REGION Network 8: End Switch
   #tmON_WaitReopenConn(IN := #tPhases.xReopenConnection, PT := T#1s);   // TON
   #tPhases.xEndSwitch := #tmON_WaitReopenConn.Q;
   IF #tmON_WaitReopenConn.Q THEN #tPhases.xReopenConnection := FALSE; END_IF;
END_REGION

REGION Network 9: - - - - - - - - Send - - - - - - - - -
END_REGION

REGION Network 10: Send Data Time Out
   #tmON_TimeoutSendData(IN := #tPhases.xRequestSend, PT := #CONST_DTIMEOUTSENDDATA_MS);   // TON
END_REGION

REGION Network 11: Request Send
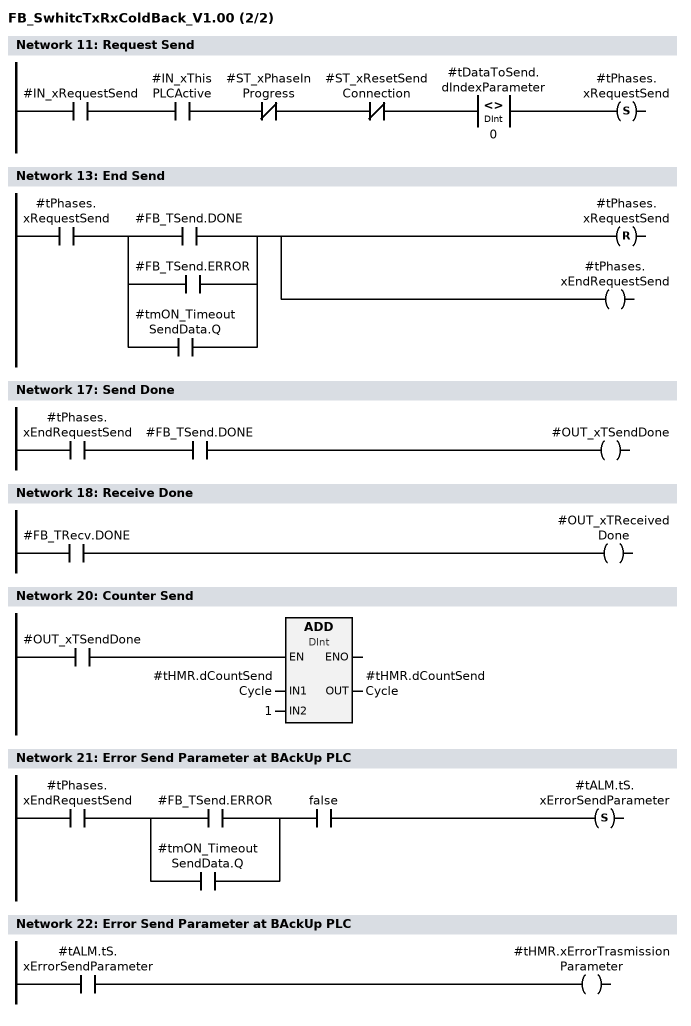
   RUNG wire#powerrail
      Contact( #IN_xRequestSend )
      Contact( #IN_xThisPLCActive )
      I_Contact( #ST_xPhaseInProgress )
      I_Contact( #ST_xResetSendConnection )
      { S7_Templates := "SrcType := DInt" } NE_Contact(in1 := #tDataToSend.dIndexParameter, in2 := 0)
      S_Coil( #tPhases.xRequestSend )
   END_RUNG
   // the same network as SCL:
   IF #IN_xRequestSend AND #IN_xThisPLCActive AND NOT #ST_xPhaseInProgress AND NOT #ST_xResetSendConnection AND (#tDataToSend.dIndexParameter <> 0) THEN
       #tPhases.xRequestSend := TRUE;
   END_IF;
END_REGION

REGION Network 12 (SCL): Send Function
       #AUX_dNumByteToSend := #tDataToSend.dByteToSend+8;//(byte for the index to send and the byte so send
   IF #tPhases.xCloseExistinConnection OR NOT #ST_xPLCActive THEN
       #FB_TSend(REQ :=FALSE,
                 CONT := FALSE,
                 LEN := #AUX_dNumByteToSend,
                 CONNECT := #AUX_tConnDataTSend,
                 DATA := #tDataToSend,
                 COM_RST := #ST_xResetSendConnection);

   ELSE
       #FB_TSend(REQ := #tPhases.xRequestSend,
                 CONT := true,
                 LEN := #AUX_dNumByteToSend,
                 CONNECT := #AUX_tConnDataTSend,
                 DATA := #tDataToSend,
                 COM_RST := #ST_xResetSendConnection);
   END_IF;
END_REGION

REGION Network 13: End Send
   RUNG wire#powerrail
      Contact( #tPhases.xRequestSend )
      wire#w1
      Contact( #FB_TSend.DONE )
      wire#w2
      R_Coil( #tPhases.xRequestSend )
   END_RUNG
   RUNG wire#w1
      Contact( #FB_TSend.ERROR )
   END_RUNG wire#w2
   RUNG wire#w1
      Contact( #tmON_TimeoutSendData.Q )
   END_RUNG wire#w2
   RUNG wire#w2
      Coil( #tPhases.xEndRequestSend )
   END_RUNG
   // the same network as SCL:
   #_w1 := #tPhases.xRequestSend AND (#FB_TSend.DONE OR #FB_TSend.ERROR OR #tmON_TimeoutSendData.Q);
   IF #_w1 THEN #tPhases.xRequestSend := FALSE; END_IF;
   #tPhases.xEndRequestSend := #_w1;
END_REGION

REGION Network 14: - - - - - - - - Recive - - - - - - - - -
END_REGION

REGION Network 15 (SCL): Recived Connection
   IF #tPhases.xCloseExistinConnection OR  #ST_xPLCActive THEN
       #FB_TRecv(EN_R := FALSE,
                 CONT := FALSE,
                 LEN := 0,
                 ADHOC:=TRUE,
                 CONNECT := #AUX_tConnDataTRecive,
                 DATA := #tDataRecived,
                 COM_RST := #ST_xResetRecvConnection);
   ELSE
       //Clean DB data recive
       FILL_BLK(IN := 0,
                COUNT := 501,
                OUT => #tDataRecived.rgbSendBuffer[0]);

       #FB_TRecv(EN_R := True,
                  CONT := True,
                  LEN := 0,
                  ADHOC:=TRUE,
                  CONNECT := #AUX_tConnDataTRecive,
                  DATA := #tDataRecived,
                  COM_RST := #ST_xResetRecvConnection);
   END_IF;
END_REGION

REGION Network 16 (SCL): Phase in progress
   GATHER(IN:=#tPhases,
          OUT=>#TMP_dwValue);

   IF #TMP_dwValue <> 0 THEN
       #ST_xPhaseInProgress := TRUE;
   ELSE
       #ST_xPhaseInProgress := FALSE;
   END_IF;
END_REGION

REGION Network 17: Send Done
   RUNG wire#powerrail
      Contact( #tPhases.xEndRequestSend )
      Contact( #FB_TSend.DONE )
      Coil( #OUT_xTSendDone )
   END_RUNG
   // the same network as SCL:
   #OUT_xTSendDone := #tPhases.xEndRequestSend AND #FB_TSend.DONE;
END_REGION

REGION Network 18: Receive Done
   RUNG wire#powerrail
      Contact( #FB_TRecv.DONE )
      Coil( #OUT_xTReceivedDone )
   END_RUNG
   // the same network as SCL:
   #OUT_xTReceivedDone := #FB_TRecv.DONE;
END_REGION

REGION Network 19: - - - - - - - -- - - HMI - - - - - - -
END_REGION

REGION Network 20: Counter Send
   RUNG wire#powerrail
      Contact( #OUT_xTSendDone )
      { S7_Templates := "SrcType := DInt" } Add(in1 := #tHMR.dCountSendCycle, in2 := 1, out => #tHMR.dCountSendCycle)
   END_RUNG
   // the same network as SCL:
   IF #OUT_xTSendDone THEN #tHMR.dCountSendCycle := #tHMR.dCountSendCycle + 1; END_IF;
END_REGION

REGION Network 21: Error Send Parameter at BAckUp PLC
   RUNG wire#powerrail
      Contact( #tPhases.xEndRequestSend )
      wire#w1
      Contact( #FB_TSend.ERROR )
      wire#w2
      Contact( false )
      S_Coil( #tALM.tS.xErrorSendParameter )
   END_RUNG
   RUNG wire#w1
      Contact( #tmON_TimeoutSendData.Q )
   END_RUNG wire#w2
   // the same network as SCL:
   IF #tPhases.xEndRequestSend AND (#FB_TSend.ERROR OR #tmON_TimeoutSendData.Q) AND false THEN
       #tALM.tS.xErrorSendParameter := TRUE;
   END_IF;
END_REGION

REGION Network 22: Error Send Parameter at BAckUp PLC
   RUNG wire#powerrail
      Contact( #tALM.tS.xErrorSendParameter )
      Coil( #tHMR.xErrorTrasmissionParameter )
   END_RUNG
   // the same network as SCL:
   #tHMR.xErrorTrasmissionParameter := #tALM.tS.xErrorSendParameter;
END_REGION
END_FUNCTION_BLOCK

FUNCTION "ExChangeParTxRx_Logic" : Void   // FC340, LAD
{ S7_Optimized_Access := 'TRUE' }
VERSION : 0.1
   VAR_INPUT
      IN_tConfDataMaster : Struct   // Configuration data master CPU
         Header : IF_CONF_Header;
         IPData : IF_CONF_v4;
         NoS : IF_CONF_NOS;
         NTP : IF_CONF_NTP;
         IP_V6 : IF_CONF_v6;
         MAC : IF_CONF_MAC;
         DNS : IF_CONF_DNS;
      END_STRUCT;
      IN_tConfDataBackup : Struct   // Configuration data backup CPU
         Header : IF_CONF_Header;
         IPData : IF_CONF_v4;
         NoS : IF_CONF_NOS;
         NTP : IF_CONF_NTP;
         IP_V6 : IF_CONF_v6;
         MAC : IF_CONF_MAC;
         DNS : IF_CONF_DNS;
      END_STRUCT;
   END_VAR
   VAR_TEMP
      TMP_x : Bool;
      TMP_dBufferPos : DInt;
      TMP_xRetValue : Int;
      IpAddress : IP_V4;
   END_VAR
BEGIN

REGION Network 1 (SCL): IP Secondary CPU
   #IpAddress.ADDR[1] := 192;
   #IpAddress.ADDR[2] := 168;
   #IpAddress.ADDR[3] := 130;
   #IpAddress.ADDR[4] := 8;
END_REGION

REGION Network 2: Call Function Swtich Send/Recive
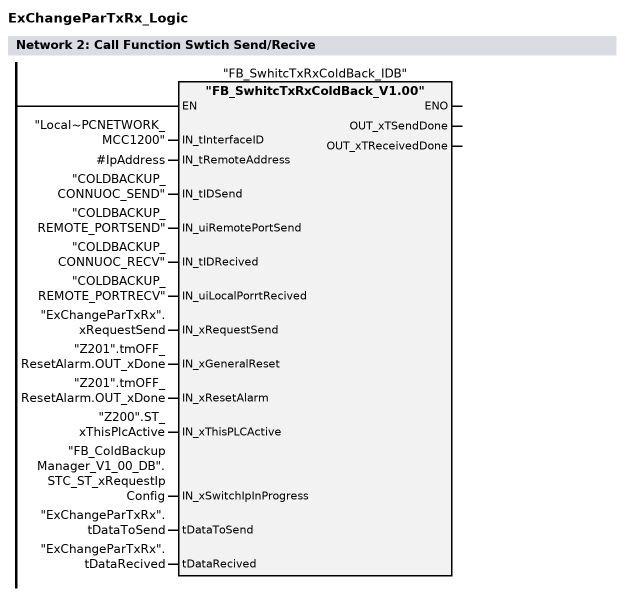
   RUNG wire#powerrail
      "FB_SwhitcTxRxColdBack_IDB"(IN_tInterfaceID := "Local~PCNETWORK_MCC1200", IN_tRemoteAddress := #IpAddress, IN_tIDSend := "COLDBACKUP_CONNUOC_SEND", IN_uiRemotePortSend := "COLDBACKUP_REMOTE_PORTSEND", IN_tIDRecived := "COLDBACKUP_CONNUOC_RECV", IN_uiLocalPorrtRecived := "COLDBACKUP_REMOTE_PORTRECV", IN_xRequestSend := "ExChangeParTxRx".xRequestSend, IN_xGeneralReset := "Z201".tmOFF_ResetAlarm.OUT_xDone, IN_xResetAlarm := "Z201".tmOFF_ResetAlarm.OUT_xDone, IN_xThisPLCActive := "Z200".ST_xThisPlcActive, IN_xSwitchIpInProgress := "FB_ColdBackupManager_V1_00_DB".STC_ST_xRequestIpConfig, tDataToSend := "ExChangeParTxRx".tDataToSend, tDataRecived := "ExChangeParTxRx".tDataRecived, OUT_xTSendDone =>, OUT_xTReceivedDone =>)
   END_RUNG
   // the same network as SCL:
   "FB_SwhitcTxRxColdBack_IDB"(IN_tInterfaceID := "Local~PCNETWORK_MCC1200",   // "FB_SwhitcTxRxColdBack_V1.00"
                           IN_tRemoteAddress := #IpAddress,
                           IN_tIDSend := "COLDBACKUP_CONNUOC_SEND",
                           IN_uiRemotePortSend := "COLDBACKUP_REMOTE_PORTSEND",
                           IN_tIDRecived := "COLDBACKUP_CONNUOC_RECV",
                           IN_uiLocalPorrtRecived := "COLDBACKUP_REMOTE_PORTRECV",
                           IN_xRequestSend := "ExChangeParTxRx".xRequestSend,
                           IN_xGeneralReset := "Z201".tmOFF_ResetAlarm.OUT_xDone,
                           IN_xResetAlarm := "Z201".tmOFF_ResetAlarm.OUT_xDone,
                           IN_xThisPLCActive := "Z200".ST_xThisPlcActive,
                           IN_xSwitchIpInProgress := "FB_ColdBackupManager_V1_00_DB".STC_ST_xRequestIpConfig,
                           tDataToSend := "ExChangeParTxRx".tDataToSend,
                           tDataRecived := "ExChangeParTxRx".tDataRecived);
END_REGION

REGION Network 3 (SCL): PLC Active Send

   IF "Z200".ST_xThisPlcActive THEN
       IF "FB_SwhitcTxRxColdBack_IDB".OUT_xTSendDone THEN
           "ExChangeParTxRx".AUX_dIndexToSend := "ExChangeParTxRx".AUX_dIndexToSend + 1;
       END_IF;

       "ExChangeParTxRx".xRequestSend := TRUE;

       CASE "ExChangeParTxRx".AUX_dIndexToSend OF
           1:  //Z200 HMW
               #TMP_dBufferPos := 0;
               #TMP_xRetValue := Serialize(SRC_VARIABLE := "DB_Z200_HMI".tHMW, DEST_ARRAY =>"ExChangeParTxRx".tDataToSend.rgbBuffer, POS := #TMP_dBufferPos);
               "ExChangeParTxRx".tDataToSend.dIndexParameter := "ExChangeParTxRx".AUX_dIndexToSend;
               "ExChangeParTxRx".tDataToSend.dNByteBuffer := #TMP_dBufferPos;

           2:  //Z200 HMR 
               #TMP_dBufferPos := 0;
               #TMP_xRetValue := Serialize(SRC_VARIABLE := "DB_Z200_HMI".tHMR, DEST_ARRAY =>"ExChangeParTxRx".tDataToSend.rgbBuffer, POS := #TMP_dBufferPos);
               "ExChangeParTxRx".tDataToSend.dIndexParameter := "ExChangeParTxRx".AUX_dIndexToSend;
               "ExChangeParTxRx".tDataToSend.dNByteBuffer := #TMP_dBufferPos;

           37:  //Z201 HMW
               #TMP_dBufferPos := 0;
               #TMP_xRetValue := Serialize(SRC_VARIABLE := "DB_Z200_HMI".tHMW, DEST_ARRAY => "ExChangeParTxRx".tDataToSend.rgbBuffer, POS := #TMP_dBufferPos);
               "ExChangeParTxRx".tDataToSend.dIndexParameter := "ExChangeParTxRx".AUX_dIndexToSend;
               "ExChangeParTxRx".tDataToSend.dNByteBuffer := #TMP_dBufferPos;

           38:  //Z201 HMR 
               #TMP_dBufferPos := 0;
               #TMP_xRetValue := Serialize(SRC_VARIABLE := "DB_Z201_HMI".tHMR, DEST_ARRAY => "ExChangeParTxRx".tDataToSend.rgbBuffer, POS := #TMP_dBufferPos);
               "ExChangeParTxRx".tDataToSend.dIndexParameter := "ExChangeParTxRx".AUX_dIndexToSend;
               "ExChangeParTxRx".tDataToSend.dNByteBuffer := #TMP_dBufferPos;

           39:  //ZUPS HMW
               #TMP_dBufferPos := 0;
               #TMP_xRetValue := Serialize(SRC_VARIABLE := "DB_ZUPS_HMI".tHMW, DEST_ARRAY => "ExChangeParTxRx".tDataToSend.rgbBuffer, POS := #TMP_dBufferPos);
               "ExChangeParTxRx".tDataToSend.dIndexParameter := "ExChangeParTxRx".AUX_dIndexToSend;
               "ExChangeParTxRx".tDataToSend.dNByteBuffer := #TMP_dBufferPos;

           40:  //ZUPS HMR 
               #TMP_dBufferPos := 0;
               #TMP_xRetValue := Serialize(SRC_VARIABLE := "DB_ZUPS_HMI".tHMR, DEST_ARRAY => "ExChangeParTxRx".tDataToSend.rgbBuffer, POS := #TMP_dBufferPos);
               "ExChangeParTxRx".tDataToSend.dIndexParameter := "ExChangeParTxRx".AUX_dIndexToSend;
               "ExChangeParTxRx".tDataToSend.dNByteBuffer := #TMP_dBufferPos;



           3:  //M201 HMW
               #TMP_dBufferPos := 0;
               #TMP_xRetValue := Serialize(SRC_VARIABLE := "FB_BD_BreakPH_V1_00_IDB".tHMW, DEST_ARRAY =>"ExChangeParTxRx".tDataToSend.rgbBuffer, POS := #TMP_dBufferPos);
               "ExChangeParTxRx".tDataToSend.dIndexParameter := "ExChangeParTxRx".AUX_dIndexToSend;
               "ExChangeParTxRx".tDataToSend.dNByteBuffer := #TMP_dBufferPos;

           4:  //M201 HMR 
               #TMP_dBufferPos := 0;
               #TMP_xRetValue := Serialize(SRC_VARIABLE := "FB_BD_BreakPH_V1_00_IDB".tHMR, DEST_ARRAY =>"ExChangeParTxRx".tDataToSend.rgbBuffer, POS := #TMP_dBufferPos);
               "ExChangeParTxRx".tDataToSend.dIndexParameter := "ExChangeParTxRx".AUX_dIndexToSend;
               "ExChangeParTxRx".tDataToSend.dNByteBuffer := #TMP_dBufferPos;

           5:  //M216 DIGITIZER HMW
               #TMP_dBufferPos := 0;
               #TMP_xRetValue := Serialize(SRC_VARIABLE := "FB_BD_DigitizerPH_V1_00_IDB".tHMW, DEST_ARRAY =>"ExChangeParTxRx".tDataToSend.rgbBuffer, POS := #TMP_dBufferPos);
               "ExChangeParTxRx".tDataToSend.dIndexParameter := "ExChangeParTxRx".AUX_dIndexToSend;
               "ExChangeParTxRx".tDataToSend.dNByteBuffer := #TMP_dBufferPos;

           6:  //M216 DIGITIZER HMR 
               #TMP_dBufferPos := 0;
               #TMP_xRetValue := Serialize(SRC_VARIABLE := "FB_BD_DigitizerPH_V1_00_IDB".tHMR, DEST_ARRAY =>"ExChangeParTxRx".tDataToSend.rgbBuffer, POS := #TMP_dBufferPos);
               "ExChangeParTxRx".tDataToSend.dIndexParameter := "ExChangeParTxRx".AUX_dIndexToSend;
               "ExChangeParTxRx".tDataToSend.dNByteBuffer := #TMP_dBufferPos;


           7:  //CrossCut 1 HMW 
               #TMP_dBufferPos := 0;
               #TMP_xRetValue := Serialize(SRC_VARIABLE := "FB_CrossCuts_1_V1_00_IDB".tHMW, DEST_ARRAY =>"ExChangeParTxRx".tDataToSend.rgbBuffer, POS := #TMP_dBufferPos);
               "ExChangeParTxRx".tDataToSend.dIndexParameter := "ExChangeParTxRx".AUX_dIndexToSend;
               "ExChangeParTxRx".tDataToSend.dNByteBuffer := #TMP_dBufferPos;

           8:  //CrossCut 1 HMR 
               #TMP_dBufferPos := 0;
               #TMP_xRetValue := Serialize(SRC_VARIABLE := "FB_CrossCuts_1_V1_00_IDB".tHMR, DEST_ARRAY =>"ExChangeParTxRx".tDataToSend.rgbBuffer, POS := #TMP_dBufferPos);
               "ExChangeParTxRx".tDataToSend.dIndexParameter := "ExChangeParTxRx".AUX_dIndexToSend;
               "ExChangeParTxRx".tDataToSend.dNByteBuffer := #TMP_dBufferPos;

           9:  //CrossCut 2 HMW 
               #TMP_dBufferPos := 0;
               #TMP_xRetValue := Serialize(SRC_VARIABLE := "FB_CrossCuts_2_V1_00_IDB".tHMW, DEST_ARRAY =>"ExChangeParTxRx".tDataToSend.rgbBuffer, POS := #TMP_dBufferPos);
               "ExChangeParTxRx".tDataToSend.dIndexParameter := "ExChangeParTxRx".AUX_dIndexToSend;
               "ExChangeParTxRx".tDataToSend.dNByteBuffer := #TMP_dBufferPos;

           10:  //CrossCut 2 HMR 
               #TMP_dBufferPos := 0;
               #TMP_xRetValue := Serialize(SRC_VARIABLE := "FB_CrossCuts_2_V1_00_IDB".tHMR, DEST_ARRAY =>"ExChangeParTxRx".tDataToSend.rgbBuffer, POS := #TMP_dBufferPos);
               "ExChangeParTxRx".tDataToSend.dIndexParameter := "ExChangeParTxRx".AUX_dIndexToSend;
               "ExChangeParTxRx".tDataToSend.dNByteBuffer := #TMP_dBufferPos;

           11:  //Digitizer 1 HMR 
               #TMP_dBufferPos := 0;
               #TMP_xRetValue := Serialize(SRC_VARIABLE := "FB_Digitizer_1_V1_00_IDB".tHMR, DEST_ARRAY =>"ExChangeParTxRx".tDataToSend.rgbBuffer, POS := #TMP_dBufferPos);
               "ExChangeParTxRx".tDataToSend.dIndexParameter := "ExChangeParTxRx".AUX_dIndexToSend;
               "ExChangeParTxRx".tDataToSend.dNByteBuffer := #TMP_dBufferPos;

           12:  //Digitizer 1 HMW 
               #TMP_dBufferPos := 0;
               #TMP_xRetValue := Serialize(SRC_VARIABLE := "FB_Digitizer_1_V1_00_IDB".tHMW, DEST_ARRAY =>"ExChangeParTxRx".tDataToSend.rgbBuffer, POS := #TMP_dBufferPos);
               "ExChangeParTxRx".tDataToSend.dIndexParameter := "ExChangeParTxRx".AUX_dIndexToSend;
               "ExChangeParTxRx".tDataToSend.dNByteBuffer := #TMP_dBufferPos;

           13:  //Digitizer 2 HMR 
               #TMP_dBufferPos := 0;
               #TMP_xRetValue := Serialize(SRC_VARIABLE := "FB_Digitizer_2_V1_00_IDB".tHMR, DEST_ARRAY =>"ExChangeParTxRx".tDataToSend.rgbBuffer, POS := #TMP_dBufferPos);
               "ExChangeParTxRx".tDataToSend.dIndexParameter := "ExChangeParTxRx".AUX_dIndexToSend;
               "ExChangeParTxRx".tDataToSend.dNByteBuffer := #TMP_dBufferPos;

           14:  //Digitizer 2 HMW 
               #TMP_dBufferPos := 0;
               #TMP_xRetValue := Serialize(SRC_VARIABLE := "FB_Digitizer_2_V1_00_IDB".tHMW, DEST_ARRAY =>"ExChangeParTxRx".tDataToSend.rgbBuffer, POS := #TMP_dBufferPos);
               "ExChangeParTxRx".tDataToSend.dIndexParameter := "ExChangeParTxRx".AUX_dIndexToSend;
               "ExChangeParTxRx".tDataToSend.dNByteBuffer := #TMP_dBufferPos;

           15:  //DigitizerManager HMR 
               #TMP_dBufferPos := 0;
               #TMP_xRetValue := Serialize(SRC_VARIABLE := "FB_DigitizerManager_V1_00_IDB".tHMR, DEST_ARRAY =>"ExChangeParTxRx".tDataToSend.rgbBuffer, POS := #TMP_dBufferPos);
               "ExChangeParTxRx".tDataToSend.dIndexParameter := "ExChangeParTxRx".AUX_dIndexToSend;
               "ExChangeParTxRx".tDataToSend.dNByteBuffer := #TMP_dBufferPos;

           16:  //DigitizerManager HMW 
               #TMP_dBufferPos := 0;
               #TMP_xRetValue := Serialize(SRC_VARIABLE := "FB_DigitizerManager_V1_00_IDB".tHMW, DEST_ARRAY =>"ExChangeParTxRx".tDataToSend.rgbBuffer, POS := #TMP_dBufferPos);
               "ExChangeParTxRx".tDataToSend.dIndexParameter := "ExChangeParTxRx".AUX_dIndexToSend;
               "ExChangeParTxRx".tDataToSend.dNByteBuffer := #TMP_dBufferPos;

           17:  //ISRA 5D HMMR
               #TMP_dBufferPos := 0;
               #TMP_xRetValue := Serialize(SRC_VARIABLE := "FB_ISRA5D_IDB".tHMR, DEST_ARRAY =>"ExChangeParTxRx".tDataToSend.rgbBuffer, POS := #TMP_dBufferPos);
               "ExChangeParTxRx".tDataToSend.dIndexParameter := "ExChangeParTxRx".AUX_dIndexToSend;
               "ExChangeParTxRx".tDataToSend.dNByteBuffer := #TMP_dBufferPos;

           18:  //ISRA 5D HMW 
               #TMP_dBufferPos := 0;
               #TMP_xRetValue := Serialize(SRC_VARIABLE := "FB_ISRA5D_IDB".tHMW, DEST_ARRAY =>"ExChangeParTxRx".tDataToSend.rgbBuffer, POS := #TMP_dBufferPos);
               "ExChangeParTxRx".tDataToSend.dIndexParameter := "ExChangeParTxRx".AUX_dIndexToSend;
               "ExChangeParTxRx".tDataToSend.dNByteBuffer := #TMP_dBufferPos;

           19:  //Man Insp HMMR
               #TMP_dBufferPos := 0;
               #TMP_xRetValue := Serialize(SRC_VARIABLE := "FB_ManInsp_V1_00_IDB".tHMR, DEST_ARRAY =>"ExChangeParTxRx".tDataToSend.rgbBuffer, POS := #TMP_dBufferPos);
               "ExChangeParTxRx".tDataToSend.dIndexParameter := "ExChangeParTxRx".AUX_dIndexToSend;
               "ExChangeParTxRx".tDataToSend.dNByteBuffer := #TMP_dBufferPos;

           20:  //Man Insp HMW 
               #TMP_dBufferPos := 0;
               #TMP_xRetValue := Serialize(SRC_VARIABLE := "FB_ManInsp_V1_00_IDB".tHMW, DEST_ARRAY =>"ExChangeParTxRx".tDataToSend.rgbBuffer, POS := #TMP_dBufferPos);
               "ExChangeParTxRx".tDataToSend.dIndexParameter := "ExChangeParTxRx".AUX_dIndexToSend;
               "ExChangeParTxRx".tDataToSend.dNByteBuffer := #TMP_dBufferPos;

           21:  //Markers HMMR
               #TMP_dBufferPos := 0;
               #TMP_xRetValue := Serialize(SRC_VARIABLE := "FB_Markers_V1.00_IDB".tHMR, DEST_ARRAY =>"ExChangeParTxRx".tDataToSend.rgbBuffer, POS := #TMP_dBufferPos);
               "ExChangeParTxRx".tDataToSend.dIndexParameter := "ExChangeParTxRx".AUX_dIndexToSend;
               "ExChangeParTxRx".tDataToSend.dNByteBuffer := #TMP_dBufferPos;

           22:  //Markers HMW 
               #TMP_dBufferPos := 0;
               #TMP_xRetValue := Serialize(SRC_VARIABLE := "FB_Markers_V1.00_IDB".tHMW, DEST_ARRAY =>"ExChangeParTxRx".tDataToSend.rgbBuffer, POS := #TMP_dBufferPos);
               "ExChangeParTxRx".tDataToSend.dIndexParameter := "ExChangeParTxRx".AUX_dIndexToSend;
               "ExChangeParTxRx".tDataToSend.dNByteBuffer := #TMP_dBufferPos;

           23:  //Oil HMMR
               #TMP_dBufferPos := 0;
               #TMP_xRetValue := Serialize(SRC_VARIABLE := "FB_Oil_V1_00_IDB".tHMR, DEST_ARRAY =>"ExChangeParTxRx".tDataToSend.rgbBuffer, POS := #TMP_dBufferPos);
               "ExChangeParTxRx".tDataToSend.dIndexParameter := "ExChangeParTxRx".AUX_dIndexToSend;
               "ExChangeParTxRx".tDataToSend.dNByteBuffer := #TMP_dBufferPos;

           24:  //Oil HMW 
               #TMP_dBufferPos := 0;
               #TMP_xRetValue := Serialize(SRC_VARIABLE := "FB_Oil_V1_00_IDB".tHMW, DEST_ARRAY =>"ExChangeParTxRx".tDataToSend.rgbBuffer, POS := #TMP_dBufferPos);
               "ExChangeParTxRx".tDataToSend.dIndexParameter := "ExChangeParTxRx".AUX_dIndexToSend;
               "ExChangeParTxRx".tDataToSend.dNByteBuffer := #TMP_dBufferPos;

           25:  //YCut 1 HMR
               #TMP_dBufferPos := 0;
               #TMP_xRetValue := Serialize(SRC_VARIABLE := "FB_YCuts1_V1_00_IDB".tHMR, DEST_ARRAY =>"ExChangeParTxRx".tDataToSend.rgbBuffer, POS := #TMP_dBufferPos);
               "ExChangeParTxRx".tDataToSend.dIndexParameter := "ExChangeParTxRx".AUX_dIndexToSend;
               "ExChangeParTxRx".tDataToSend.dNByteBuffer := #TMP_dBufferPos;

           26:  //YCut 1 HMW
               #TMP_dBufferPos := 0;
               #TMP_xRetValue := Serialize(SRC_VARIABLE := "FB_YCuts1_V1_00_IDB".tHMW, DEST_ARRAY =>"ExChangeParTxRx".tDataToSend.rgbBuffer, POS := #TMP_dBufferPos);
               "ExChangeParTxRx".tDataToSend.dIndexParameter := "ExChangeParTxRx".AUX_dIndexToSend;
               "ExChangeParTxRx".tDataToSend.dNByteBuffer := #TMP_dBufferPos;

           27:  //YCut 2 HMR
               #TMP_dBufferPos := 0;
               #TMP_xRetValue := Serialize(SRC_VARIABLE := "FB_YCuts2_V1_00_IDB".tHMR, DEST_ARRAY =>"ExChangeParTxRx".tDataToSend.rgbBuffer, POS := #TMP_dBufferPos);
               "ExChangeParTxRx".tDataToSend.dIndexParameter := "ExChangeParTxRx".AUX_dIndexToSend;
               "ExChangeParTxRx".tDataToSend.dNByteBuffer := #TMP_dBufferPos;

           28:  //YCut 2 HMW
               #TMP_dBufferPos := 0;
               #TMP_xRetValue := Serialize(SRC_VARIABLE := "FB_YCuts2_V1_00_IDB".tHMW, DEST_ARRAY =>"ExChangeParTxRx".tDataToSend.rgbBuffer, POS := #TMP_dBufferPos);
               "ExChangeParTxRx".tDataToSend.dIndexParameter := "ExChangeParTxRx".AUX_dIndexToSend;
               "ExChangeParTxRx".tDataToSend.dNByteBuffer := #TMP_dBufferPos;

           29:  //OPT Manager HMR
               #TMP_dBufferPos := 0;
               #TMP_xRetValue := Serialize(SRC_VARIABLE := "FB_OptManager_V1_00_IDB".tHMR, DEST_ARRAY =>"ExChangeParTxRx".tDataToSend.rgbBuffer, POS := #TMP_dBufferPos);
               "ExChangeParTxRx".tDataToSend.dIndexParameter := "ExChangeParTxRx".AUX_dIndexToSend;
               "ExChangeParTxRx".tDataToSend.dNByteBuffer := #TMP_dBufferPos;

           30:  //OPT Manager HMW
               #TMP_dBufferPos := 0;
               #TMP_xRetValue := Serialize(SRC_VARIABLE := "FB_OptManager_V1_00_IDB".tHMW, DEST_ARRAY =>"ExChangeParTxRx".tDataToSend.rgbBuffer, POS := #TMP_dBufferPos);
               "ExChangeParTxRx".tDataToSend.dIndexParameter := "ExChangeParTxRx".AUX_dIndexToSend;
               "ExChangeParTxRx".tDataToSend.dNByteBuffer := #TMP_dBufferPos;

           31:  //Snaproll HMR
               #TMP_dBufferPos := 0;
               #TMP_xRetValue := Serialize(SRC_VARIABLE := "FB_Snaproll_V1_00_IDB".tHMR, DEST_ARRAY => "ExChangeParTxRx".tDataToSend.rgbBuffer, POS := #TMP_dBufferPos);
               "ExChangeParTxRx".tDataToSend.dIndexParameter := "ExChangeParTxRx".AUX_dIndexToSend;
               "ExChangeParTxRx".tDataToSend.dNByteBuffer := #TMP_dBufferPos;

           32:  //Snaproll HMW
               #TMP_dBufferPos := 0;
               #TMP_xRetValue := Serialize(SRC_VARIABLE := "FB_Snaproll_V1_00_IDB".tHMW, DEST_ARRAY => "ExChangeParTxRx".tDataToSend.rgbBuffer, POS := #TMP_dBufferPos);
               "ExChangeParTxRx".tDataToSend.dIndexParameter := "ExChangeParTxRx".AUX_dIndexToSend;
               "ExChangeParTxRx".tDataToSend.dNByteBuffer := #TMP_dBufferPos;

           33:  //LehrSpeed HMR
               #TMP_dBufferPos := 0;
               #TMP_xRetValue := Serialize(SRC_VARIABLE := "FB_LehrSpeed_IDB".tHMR, DEST_ARRAY => "ExChangeParTxRx".tDataToSend.rgbBuffer, POS := #TMP_dBufferPos);
               "ExChangeParTxRx".tDataToSend.dIndexParameter := "ExChangeParTxRx".AUX_dIndexToSend;
               "ExChangeParTxRx".tDataToSend.dNByteBuffer := #TMP_dBufferPos;

           34:  //LehrSpeed HMW
               #TMP_dBufferPos := 0;
               #TMP_xRetValue := Serialize(SRC_VARIABLE := "FB_LehrSpeed_IDB".tHMW, DEST_ARRAY => "ExChangeParTxRx".tDataToSend.rgbBuffer, POS := #TMP_dBufferPos);
               "ExChangeParTxRx".tDataToSend.dIndexParameter := "ExChangeParTxRx".AUX_dIndexToSend;
               "ExChangeParTxRx".tDataToSend.dNByteBuffer := #TMP_dBufferPos;

           35:  //Wander camera HMR
               #TMP_dBufferPos := 0;
               #TMP_xRetValue := Serialize(SRC_VARIABLE := "FB_WanderCamera_V1_00_IDB".tHMR, DEST_ARRAY => "ExChangeParTxRx".tDataToSend.rgbBuffer, POS := #TMP_dBufferPos);
               "ExChangeParTxRx".tDataToSend.dIndexParameter := "ExChangeParTxRx".AUX_dIndexToSend;
               "ExChangeParTxRx".tDataToSend.dNByteBuffer := #TMP_dBufferPos;

           36:  //Wander camera HMW
               #TMP_dBufferPos := 0;
               #TMP_xRetValue := Serialize(SRC_VARIABLE := "FB_WanderCamera_V1_00_IDB".tHMW, DEST_ARRAY => "ExChangeParTxRx".tDataToSend.rgbBuffer, POS := #TMP_dBufferPos);
               "ExChangeParTxRx".tDataToSend.dIndexParameter := "ExChangeParTxRx".AUX_dIndexToSend;
               "ExChangeParTxRx".tDataToSend.dNByteBuffer := #TMP_dBufferPos;


           ELSE  // Statement section ELSE
               "ExChangeParTxRx".AUX_dIndexToSend := 1;
               "ExChangeParTxRx".xRequestSend := FALSE;
       END_CASE;

   ELSE
       "ExChangeParTxRx".xRequestSend:=FALSE;
   END_IF;
END_REGION

REGION Network 4 (SCL): PLC not Active Recived Conversion

   IF NOT "Z200".ST_xThisPlcActive THEN
       IF "FB_SwhitcTxRxColdBack_IDB".OUT_xTReceivedDone THEN
           CASE "ExChangeParTxRx".tDataRecived.dIndexParameter OF

               1:  //Z200 HMW
                   #TMP_dBufferPos := 0;
                   #TMP_xRetValue := Deserialize(SRC_ARRAY := "ExChangeParTxRx".tDataRecived.rgbBuffer, DEST_VARIABLE => "DB_Z200_HMI".tHMW, POS := #TMP_dBufferPos);

               2:  //Z200 HMR 
                   #TMP_dBufferPos := 0;
                   #TMP_xRetValue := Deserialize(SRC_ARRAY := "ExChangeParTxRx".tDataRecived.rgbBuffer, DEST_VARIABLE => "DB_Z200_HMI".tHMR, POS := #TMP_dBufferPos);

               37:  //Z201 HMW
                   #TMP_dBufferPos := 0;
                   #TMP_xRetValue := Deserialize(SRC_ARRAY := "ExChangeParTxRx".tDataRecived.rgbBuffer, DEST_VARIABLE => "DB_Z201_HMI".tHMW, POS := #TMP_dBufferPos);

               38:  //Z201 HMR 
                   #TMP_dBufferPos := 0;
                   #TMP_xRetValue := Deserialize(SRC_ARRAY := "ExChangeParTxRx".tDataRecived.rgbBuffer, DEST_VARIABLE => "DB_Z201_HMI".tHMR, POS := #TMP_dBufferPos);

               39:  //ZUPS HMW
                   #TMP_dBufferPos := 0;
                   #TMP_xRetValue := Deserialize(SRC_ARRAY := "ExChangeParTxRx".tDataRecived.rgbBuffer, DEST_VARIABLE => "DB_ZUPS_HMI".tHMW, POS := #TMP_dBufferPos);

               40:  //Z2UPS HMR 
                   #TMP_dBufferPos := 0;
                   #TMP_xRetValue := Deserialize(SRC_ARRAY := "ExChangeParTxRx".tDataRecived.rgbBuffer, DEST_VARIABLE => "DB_ZUPS_HMI".tHMR, POS := #TMP_dBufferPos);

               3:  //M201 HMW
                   #TMP_dBufferPos := 0;
                   #TMP_xRetValue := Deserialize(SRC_ARRAY := "ExChangeParTxRx".tDataRecived.rgbBuffer, DEST_VARIABLE => "FB_BD_BreakPH_V1_00_IDB".tHMW, POS := #TMP_dBufferPos);

               4:  //M201 HMR 
                   #TMP_dBufferPos := 0;
                   #TMP_xRetValue := Deserialize(SRC_ARRAY := "ExChangeParTxRx".tDataRecived.rgbBuffer, DEST_VARIABLE => "FB_BD_BreakPH_V1_00_IDB".tHMR, POS := #TMP_dBufferPos);

               5:  //M216 Digitizer HMW
                   #TMP_dBufferPos := 0;
                   #TMP_xRetValue := Deserialize(SRC_ARRAY := "ExChangeParTxRx".tDataRecived.rgbBuffer, DEST_VARIABLE => "FB_BD_DigitizerPH_V1_00_IDB".tHMW, POS := #TMP_dBufferPos);

               6:  //M216 Digitizer HMR 
                   #TMP_dBufferPos := 0;
                   #TMP_xRetValue := Deserialize(SRC_ARRAY := "ExChangeParTxRx".tDataRecived.rgbBuffer, DEST_VARIABLE => "FB_BD_DigitizerPH_V1_00_IDB".tHMR, POS := #TMP_dBufferPos);

               7:  //CrossCut 1 HMW 
                   #TMP_dBufferPos := 0;
                   #TMP_xRetValue := Deserialize(SRC_ARRAY := "ExChangeParTxRx".tDataRecived.rgbBuffer, DEST_VARIABLE => "FB_CrossCuts_1_V1_00_IDB".tHMW, POS := #TMP_dBufferPos);

               8:  //CrossCut 1 HMR 
                   #TMP_dBufferPos := 0;
                   #TMP_xRetValue := Deserialize(SRC_ARRAY := "ExChangeParTxRx".tDataRecived.rgbBuffer, DEST_VARIABLE => "FB_CrossCuts_1_V1_00_IDB".tHMR, POS := #TMP_dBufferPos);

               9:  //CrossCut 2 HMW 
                   #TMP_dBufferPos := 0;
                   #TMP_xRetValue := Deserialize(SRC_ARRAY := "ExChangeParTxRx".tDataRecived.rgbBuffer, DEST_VARIABLE => "FB_CrossCuts_2_V1_00_IDB".tHMW, POS := #TMP_dBufferPos);

               10:  //CrossCut 2 HMR 
                   #TMP_dBufferPos := 0;
                   #TMP_xRetValue := Deserialize(SRC_ARRAY := "ExChangeParTxRx".tDataRecived.rgbBuffer, DEST_VARIABLE => "FB_CrossCuts_2_V1_00_IDB".tHMR, POS := #TMP_dBufferPos);

               11:  //Digitizer 1 HMR 
                   #TMP_dBufferPos := 0;
                   #TMP_xRetValue := Deserialize(SRC_ARRAY := "ExChangeParTxRx".tDataRecived.rgbBuffer, DEST_VARIABLE => "FB_Digitizer_1_V1_00_IDB".tHMR, POS := #TMP_dBufferPos);

               12:  //Digitizer 1 HMW 
                   #TMP_dBufferPos := 0;
                   #TMP_xRetValue := Deserialize(SRC_ARRAY := "ExChangeParTxRx".tDataRecived.rgbBuffer, DEST_VARIABLE => "FB_Digitizer_1_V1_00_IDB".tHMW, POS := #TMP_dBufferPos);

               13:  //Digitizer 2 HMR 
                   #TMP_dBufferPos := 0;
                   #TMP_xRetValue := Deserialize(SRC_ARRAY := "ExChangeParTxRx".tDataRecived.rgbBuffer, DEST_VARIABLE => "FB_Digitizer_2_V1_00_IDB".tHMR, POS := #TMP_dBufferPos);

               14:  //Digitizer 2 HMW 
                   #TMP_dBufferPos := 0;
                   #TMP_xRetValue := Deserialize(SRC_ARRAY := "ExChangeParTxRx".tDataRecived.rgbBuffer, DEST_VARIABLE => "FB_Digitizer_2_V1_00_IDB".tHMW, POS := #TMP_dBufferPos);

               15:  //DigitizerManager HMR 
                   #TMP_dBufferPos := 0;
                   #TMP_xRetValue := Deserialize(SRC_ARRAY := "ExChangeParTxRx".tDataRecived.rgbBuffer, DEST_VARIABLE => "FB_DigitizerManager_V1_00_IDB".tHMR, POS := #TMP_dBufferPos);

               16:  //DigitizerManager HMW 
                   #TMP_dBufferPos := 0;
                   #TMP_xRetValue := Deserialize(SRC_ARRAY := "ExChangeParTxRx".tDataRecived.rgbBuffer, DEST_VARIABLE => "FB_DigitizerManager_V1_00_IDB".tHMW, POS := #TMP_dBufferPos);

               17:  //ISRA 5D HMMR
                   #TMP_dBufferPos := 0;
                   #TMP_xRetValue := Deserialize(SRC_ARRAY := "ExChangeParTxRx".tDataRecived.rgbBuffer, DEST_VARIABLE => "FB_ISRA5D_IDB".tHMR, POS := #TMP_dBufferPos);

               18:  //ISRA 5D HMW 
                   #TMP_dBufferPos := 0;
                   #TMP_xRetValue := Deserialize(SRC_ARRAY := "ExChangeParTxRx".tDataRecived.rgbBuffer, DEST_VARIABLE => "FB_ISRA5D_IDB".tHMW, POS := #TMP_dBufferPos);

               19:  //Man Insp HMMR
                   #TMP_dBufferPos := 0;
                   #TMP_xRetValue := Deserialize(SRC_ARRAY := "ExChangeParTxRx".tDataRecived.rgbBuffer, DEST_VARIABLE => "FB_ManInsp_V1_00_IDB".tHMR, POS := #TMP_dBufferPos);

               20:  //Man Insp HMW 
                   #TMP_dBufferPos := 0;
                   #TMP_xRetValue := Deserialize(SRC_ARRAY := "ExChangeParTxRx".tDataRecived.rgbBuffer, DEST_VARIABLE => "FB_ManInsp_V1_00_IDB".tHMW, POS := #TMP_dBufferPos);

               21:  //Markers HMMR
                   #TMP_dBufferPos := 0;
                   #TMP_xRetValue := Deserialize(SRC_ARRAY := "ExChangeParTxRx".tDataRecived.rgbBuffer, DEST_VARIABLE => "FB_Markers_V1.00_IDB".tHMR, POS := #TMP_dBufferPos);

               22:  //Markers HMW 
                   #TMP_dBufferPos := 0;
                   #TMP_xRetValue := Deserialize(SRC_ARRAY := "ExChangeParTxRx".tDataRecived.rgbBuffer, DEST_VARIABLE => "FB_Markers_V1.00_IDB".tHMW , POS := #TMP_dBufferPos);

               23:  //Oil HMMR
                   #TMP_dBufferPos := 0;
                   #TMP_xRetValue := Deserialize(SRC_ARRAY := "ExChangeParTxRx".tDataRecived.rgbBuffer, DEST_VARIABLE => "FB_Oil_V1_00_IDB".tHMR, POS := #TMP_dBufferPos);

               24:  //Oil HMW 
                   #TMP_dBufferPos := 0;
                   #TMP_xRetValue := Deserialize(SRC_ARRAY := "ExChangeParTxRx".tDataRecived.rgbBuffer, DEST_VARIABLE => "FB_Oil_V1_00_IDB".tHMW, POS := #TMP_dBufferPos);

               25:  //YCut 1 HMR
                   #TMP_dBufferPos := 0;
                   #TMP_xRetValue := Deserialize(SRC_ARRAY := "ExChangeParTxRx".tDataRecived.rgbBuffer, DEST_VARIABLE => "FB_YCuts1_V1_00_IDB".tHMR, POS := #TMP_dBufferPos);

               26:  //YCut 1 HMW
                   #TMP_dBufferPos := 0;
                   #TMP_xRetValue := Deserialize(SRC_ARRAY := "ExChangeParTxRx".tDataRecived.rgbBuffer, DEST_VARIABLE => "FB_YCuts1_V1_00_IDB".tHMW, POS := #TMP_dBufferPos);

               27:  //YCut 2 HMR
                   #TMP_dBufferPos := 0;
                   #TMP_xRetValue := Deserialize(SRC_ARRAY := "ExChangeParTxRx".tDataRecived.rgbBuffer, DEST_VARIABLE => "FB_YCuts2_V1_00_IDB".tHMR, POS := #TMP_dBufferPos);

               28:  //YCut 2 HMW
                   #TMP_dBufferPos := 0;
                   #TMP_xRetValue := Deserialize(SRC_ARRAY := "ExChangeParTxRx".tDataRecived.rgbBuffer, DEST_VARIABLE => "FB_YCuts2_V1_00_IDB".tHMW, POS := #TMP_dBufferPos);

               29:  //OPT Manager HMR
                   #TMP_dBufferPos := 0;
                   #TMP_xRetValue := Deserialize(SRC_ARRAY := "ExChangeParTxRx".tDataRecived.rgbBuffer, DEST_VARIABLE => "FB_OptManager_V1_00_IDB".tHMR, POS := #TMP_dBufferPos);

               30:  //OPT Manager HMW
                   #TMP_dBufferPos := 0;
                   #TMP_xRetValue := Deserialize(SRC_ARRAY := "ExChangeParTxRx".tDataRecived.rgbBuffer, DEST_VARIABLE => "FB_OptManager_V1_00_IDB".tHMW, POS := #TMP_dBufferPos);

               31:  //Snaproll HMR
                   #TMP_dBufferPos := 0;
                   #TMP_xRetValue := Deserialize(SRC_ARRAY := "ExChangeParTxRx".tDataRecived.rgbBuffer, DEST_VARIABLE => "FB_Snaproll_V1_00_IDB".tHMR, POS := #TMP_dBufferPos);

               32:  //Snaproll HMW
                   #TMP_dBufferPos := 0;
                   #TMP_xRetValue := Deserialize(SRC_ARRAY := "ExChangeParTxRx".tDataRecived.rgbBuffer, DEST_VARIABLE => "FB_Snaproll_V1_00_IDB".tHMW, POS := #TMP_dBufferPos);

               33:  //LehrSpeed HMR
                   #TMP_dBufferPos := 0;
                   #TMP_xRetValue := Deserialize(SRC_ARRAY := "ExChangeParTxRx".tDataRecived.rgbBuffer, DEST_VARIABLE => "FB_LehrSpeed_IDB".tHMR, POS := #TMP_dBufferPos);

               34:  //LehrSpeed HMW
                   #TMP_dBufferPos := 0;
                   #TMP_xRetValue := Deserialize(SRC_ARRAY := "ExChangeParTxRx".tDataRecived.rgbBuffer, DEST_VARIABLE => "FB_LehrSpeed_IDB".tHMW, POS := #TMP_dBufferPos);

               35:  //Wander camera HMR
                   #TMP_dBufferPos := 0;
                   #TMP_xRetValue := Deserialize(SRC_ARRAY := "ExChangeParTxRx".tDataRecived.rgbBuffer, DEST_VARIABLE => "FB_WanderCamera_V1_00_IDB".tHMR, POS := #TMP_dBufferPos);

               36:  //Wander camera HMW
                   #TMP_dBufferPos := 0;
                   #TMP_xRetValue := Deserialize(SRC_ARRAY := "ExChangeParTxRx".tDataRecived.rgbBuffer, DEST_VARIABLE => "FB_WanderCamera_V1_00_IDB".tHMW, POS := #TMP_dBufferPos);

               ELSE  // Statement section ELSE
                   "ExChangeParTxRx".AUX_dIndexToSend := 1;
                   "ExChangeParTxRx".xRequestSend := FALSE;
           END_CASE;
       END_IF;
   END_IF;
END_REGION
END_FUNCTION

// folder: 03_Programs_Logics/MCC1200/16_Ribbon

FUNCTION_BLOCK "FB_TrackRibbon_V1.00"   // FB19, LAD
TITLE = Tracking defects
{ S7_Optimized_Access := 'TRUE' }
VERSION : 0.1
   VAR_INPUT
      IN_xFaultsEnabled : Bool;   // Faults enabled
      IN_xCycleON : Bool;   // Zone is in cycle
      IN_xGeneralReset : Bool;   // General reset
      IN_xFaultsReset : Bool;   // Reset alarms
   END_VAR
   VAR_IN_OUT
      INO_tEncoder : "UDT_Encoder";   // Encoder data
      INO_tOBInit : "GP_OB_Initialize";
      INO_tRibbon : "UDT_RibbonData";
      INO_xRibbonBufferFull : Bool;   // Ribbon buffer full
      INO_xBreakBufferFull : Bool := false;   // Break buffer full
   END_VAR
   VAR
      OSR_xGeneralReset : Bool;   // OSR.General reset
      AUX_tEmptyGlassDataSingle : "UDT_RibbonData_GlassData_SingleData";   // Empty glass data single
      AUX_tEmptyBreakDataSingle : "UDT_RibbonData_GlassBreak_SingleBreak";   // Empty break data single
      AUX_rgtLastUpdData : Array[0.."DMAXGLASSDATAMACHINE_IND"] of "UDT_RibbonData_GlassData_SingleData";   // Last updated glass data machine
      AUX_rgtLastUpdBreak : Array[0.."DMAXGLASSDATAMACHINE_IND"] of "UDT_RibbonData_GlassBreak_SingleBreak";   // Last updated break data machine
   END_VAR
   VAR_TEMP
      TMP_xOSGeneralReset : Bool;
      TMP_dIndex : DInt;
      TMP_dIndex2nd : DInt;
      TMP_dNextTail : DInt;
      TMP_dValue_cmm : DInt;
      TMP_dNextHead : DInt;
      TMP_dSourceIndex : DInt;
      TMP_dBreakMachIndex : DInt;
      TMP_xGlassBreak : Bool;
   END_VAR
   VAR CONSTANT
      CONST_DTHRDELRIBBON_CMM : DInt := 200000;   // Delete ribbon data threshold [mm/100]
      CONST_DTHRDELBREAK_CMM : DInt := 200000;   // Delete glass break threshold [mm/100]
      CONST_DSAFETYTHR_CMM : DInt := 100000;   // Safety threshold value [mm/100]
   END_VAR
   VAR_TEMP   // added for the SCL form of the ladder/FBD networks
      _w1 : Bool;
   END_VAR
BEGIN

REGION Network 1: General reset
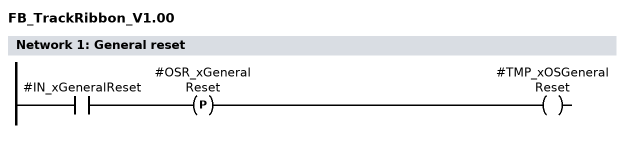
   RUNG wire#powerrail
      Contact( #IN_xGeneralReset )
      P_Trig( #OSR_xGeneralReset )
      Coil( #TMP_xOSGeneralReset )
   END_RUNG
   // the same network as SCL:
   #_w1 := #IN_xGeneralReset AND NOT #OSR_xGeneralReset;   // rising edge
   #OSR_xGeneralReset := #IN_xGeneralReset;
   #TMP_xOSGeneralReset := #_w1;
END_REGION

REGION Network 2 (SCL): Reset all the buffers
   IF #TMP_xOSGeneralReset THEN

       FOR #TMP_dIndex := 0 TO "DMAXGLASSDATAMACHINE_IND" DO

           #INO_tRibbon.rgtGlassData[#TMP_dIndex].dBufferHead := -1;
           #INO_tRibbon.rgtGlassData[#TMP_dIndex].dBufferTail := -1;
           #INO_tRibbon.rgtGlassData[#TMP_dIndex].dLastInsertEncCount_cmm := 0;

           #INO_tRibbon.rgtGlassDataUpdate[#TMP_dIndex].xUpdateRequest := FALSE;
           #AUX_rgtLastUpdData[#TMP_dIndex] := #AUX_tEmptyGlassDataSingle;

           FOR #TMP_dIndex2nd := 0 TO "DMAXGLASSDATASECTORS_IND" DO

               #INO_tRibbon.rgtGlassData[#TMP_dIndex].rgtBuffer[#TMP_dIndex2nd] := #AUX_tEmptyGlassDataSingle;

           END_FOR;        

           #INO_tRibbon.rgtGlassData[#TMP_dIndex].tLastDataBuffer := #AUX_tEmptyGlassDataSingle;

       END_FOR;

       FOR #TMP_dIndex := 0 TO "DMAXGLASSBREAKMACHINE_IND" DO

           #INO_tRibbon.rgtGlassBreak[#TMP_dIndex].dBufferHead := -1;
           #INO_tRibbon.rgtGlassBreak[#TMP_dIndex].dBufferTail := -1;
           #INO_tRibbon.rgtGlassBreak[#TMP_dIndex].dLastInsertEncCount_cmm := 0;

           #INO_tRibbon.rgtGlassBreakUpdate[#TMP_dIndex].xUpdateRequest := FALSE;
           #AUX_rgtLastUpdBreak[#TMP_dIndex] := #AUX_tEmptyBreakDataSingle;

           FOR #TMP_dIndex2nd := 0 TO "DMAXGLASSBREAKSECTORS_IND" DO

               #INO_tRibbon.rgtGlassBreak[#TMP_dIndex].rgtBuffer[#TMP_dIndex2nd] := #AUX_tEmptyBreakDataSingle;

           END_FOR;

           #INO_tRibbon.rgtGlassBreak[#TMP_dIndex].tLastDataBuffer := #AUX_tEmptyBreakDataSingle;

       END_FOR;

       FOR #TMP_dIndex := 0 TO "DMAXGLASSBREAKREQUEST_IND" DO
           #INO_tRibbon.rgtGlassBreakRequest[#TMP_dIndex].IN_dDistanceSnaproll_cmm := 0;
           #INO_tRibbon.rgtGlassBreakRequest[#TMP_dIndex].IN_dDownstreamOffset_cmm := 0;
           #INO_tRibbon.rgtGlassBreakRequest[#TMP_dIndex].IN_dUpstreamOffset_cmm := 0;
           #INO_tRibbon.rgtGlassBreakRequest[#TMP_dIndex].IN_xRequestGlassBreak := FALSE;
           #INO_tRibbon.rgtGlassBreakRequest[#TMP_dIndex].OUT_xGlassBreak := FALSE;
       END_FOR;

       FOR #TMP_dIndex := 0 TO "DMAXGLASSDATAREQUEST_IND" DO
           #INO_tRibbon.rgtGlassDataRequest[#TMP_dIndex].IN_dDistanceSnaproll_cmm := 0;
           #INO_tRibbon.rgtGlassDataRequest[#TMP_dIndex].IN_dSourceIndex := 0;
           #INO_tRibbon.rgtGlassDataRequest[#TMP_dIndex].IN_xRequestGlassData := 0;
           #INO_tRibbon.rgtGlassDataRequest[#TMP_dIndex].OUT_dGrossWander_cmm := 0;
           #INO_tRibbon.rgtGlassDataRequest[#TMP_dIndex].OUT_dGrossWidth_cmm := 0;
           #INO_tRibbon.rgtGlassDataRequest[#TMP_dIndex].OUT_dNetWander_cmm := 0;
           #INO_tRibbon.rgtGlassDataRequest[#TMP_dIndex].OUT_dNetWidth_cmm := 0;
       END_FOR;

       RETURN;

   END_IF;
END_REGION

REGION Network 3 (SCL): Delete ribbon data on buffer after position
   FOR #TMP_dIndex := 0 TO "DMAXGLASSDATAMACHINE_IND" DO 


       WHILE (#INO_tRibbon.rgtGlassData[#TMP_dIndex].dBufferTail <> #INO_tRibbon.rgtGlassData[#TMP_dIndex].dBufferHead)                                                      
                                                           AND (#INO_tRibbon.rgtGlassData[#TMP_dIndex].dBufferHead <> -1) DO

           IF (#INO_tRibbon.rgtGlassData[#TMP_dIndex].dBufferTail + 1) >= "DMAXGLASSDATASECTORS" THEN
               #TMP_dNextTail := 0;
           ELSE
               #TMP_dNextTail := #INO_tRibbon.rgtGlassData[#TMP_dIndex].dBufferTail + 1;
           END_IF;

           #TMP_dValue_cmm := #INO_tEncoder.dActualEncoderCounter_cmm - #INO_tRibbon.rgtGlassData[#TMP_dIndex].rgtBuffer[#TMP_dNextTail].dEncoderValue_cmm;

           IF (#TMP_dValue_cmm > #CONST_DTHRDELRIBBON_CMM) THEN

               #INO_tRibbon.rgtGlassData[#TMP_dIndex].tLastDataBuffer := #INO_tRibbon.rgtGlassData[#TMP_dIndex].rgtBuffer[#TMP_dNextTail];
               #INO_tRibbon.rgtGlassData[#TMP_dIndex].rgtBuffer[#TMP_dNextTail] := #AUX_tEmptyGlassDataSingle;

               #INO_tRibbon.rgtGlassData[#TMP_dIndex].tLastDataBuffer.xUpdateDataBPSA := TRUE;
               #INO_tRibbon.rgtGlassData[#TMP_dIndex].tLastDataBuffer.xUpdateDataBPSB := TRUE;

               #INO_tRibbon.rgtGlassData[#TMP_dIndex].dBufferTail := #TMP_dNextTail;

           ELSE

               EXIT; //Exit the while

           END_IF;    

       END_WHILE;    

   END_FOR;
END_REGION

REGION Network 4 (SCL): Delete break data on buffer after position
   FOR #TMP_dIndex := 0 TO "DMAXGLASSBREAKMACHINE_IND" DO

       WHILE (#INO_tRibbon.rgtGlassBreak[#TMP_dIndex].dBufferTail <> #INO_tRibbon.rgtGlassBreak[#TMP_dIndex].dBufferHead)
                                                       AND (#INO_tRibbon.rgtGlassBreak[#TMP_dIndex].dBufferHead <> -1) DO

           IF (#INO_tRibbon.rgtGlassBreak[#TMP_dIndex].dBufferTail + 1) >= "DMAXGLASSBREAKSECTORS" THEN
               #TMP_dNextTail := 0;
           ELSE
               #TMP_dNextTail := #INO_tRibbon.rgtGlassBreak[#TMP_dIndex].dBufferTail + 1;
           END_IF;

           #TMP_dValue_cmm := #INO_tEncoder.dActualEncoderCounter_cmm - #INO_tRibbon.rgtGlassBreak[#TMP_dIndex].rgtBuffer[#TMP_dNextTail].dEncoderValue_cmm;


           IF (#TMP_dValue_cmm > #CONST_DTHRDELBREAK_CMM) THEN

               #INO_tRibbon.rgtGlassBreak[#TMP_dIndex].tLastDataBuffer := #INO_tRibbon.rgtGlassBreak[#TMP_dIndex].rgtBuffer[#TMP_dNextTail];
               #INO_tRibbon.rgtGlassBreak[#TMP_dIndex].rgtBuffer[#TMP_dNextTail] := #AUX_tEmptyBreakDataSingle;

               #INO_tRibbon.rgtGlassBreak[#TMP_dIndex].dBufferTail := #TMP_dNextTail;

           ELSE

               EXIT; //Exit the while

           END_IF;

       END_WHILE;

   END_FOR;
END_REGION

REGION Network 5 (SCL): Insert the new position glass data position or update the last one
   FOR #TMP_dIndex := 0 TO #INO_tRibbon.dActualNumberGlassDataMachine - 1 DO

       //New position from external device, 
       IF (#INO_tRibbon.rgtGlassDataUpdate[#TMP_dIndex].xUpdateRequest) THEN

           //Increment the index head
           IF (#INO_tRibbon.rgtGlassData[#TMP_dIndex].dBufferHead + 1) >= "DMAXGLASSDATASECTORS" THEN
               #TMP_dNextHead := 0;
           ELSE
               #TMP_dNextHead := #INO_tRibbon.rgtGlassData[#TMP_dIndex].dBufferHead + 1;
           END_IF;

           //Check if the buffer is full
           IF (#TMP_dNextHead = #INO_tRibbon.rgtGlassData[#TMP_dIndex].dBufferTail) AND (#INO_tRibbon.rgtGlassData[#TMP_dIndex].dBufferHead <> -1) THEN
               EXIT;
           END_IF; 

           #INO_tRibbon.rgtGlassData[#TMP_dIndex].rgtBuffer[#TMP_dNextHead].dEncoderValue_cmm := #INO_tEncoder.dActualEncoderCounter_cmm + #INO_tRibbon.rgtGlassData[#TMP_dIndex].dDistSnapRoll_cmm;

           #INO_tRibbon.rgtGlassData[#TMP_dIndex].rgtBuffer[#TMP_dNextHead].dGrossWidth_cmm := #INO_tRibbon.rgtGlassDataUpdate[#TMP_dIndex].tData.dGrossWidth_cmm;
           #INO_tRibbon.rgtGlassData[#TMP_dIndex].rgtBuffer[#TMP_dNextHead].dNetWidth_cmm := #INO_tRibbon.rgtGlassDataUpdate[#TMP_dIndex].tData.dNetWidth_cmm;
           #INO_tRibbon.rgtGlassData[#TMP_dIndex].rgtBuffer[#TMP_dNextHead].dGrossWander_cmm := #INO_tRibbon.rgtGlassDataUpdate[#TMP_dIndex].tData.dGrossWander_cmm;
           #INO_tRibbon.rgtGlassData[#TMP_dIndex].rgtBuffer[#TMP_dNextHead].dNetWander_cmm := #INO_tRibbon.rgtGlassDataUpdate[#TMP_dIndex].tData.dNetWander_cmm;

           #INO_tRibbon.rgtGlassData[#TMP_dIndex].dLastInsertEncCount_cmm := #INO_tRibbon.rgtGlassData[#TMP_dIndex].rgtBuffer[#TMP_dNextHead].dEncoderValue_cmm;
           #INO_tRibbon.rgtGlassData[#TMP_dIndex].rgtBuffer[#TMP_dNextHead].xUpdateDataBPSA := TRUE;
           #INO_tRibbon.rgtGlassData[#TMP_dIndex].rgtBuffer[#TMP_dNextHead].xUpdateDataBPSB := TRUE;
           #INO_tRibbon.rgtGlassData[#TMP_dIndex].rgtBuffer[#TMP_dNextHead].xDataPresent := TRUE;


           #INO_tRibbon.rgtGlassData[#TMP_dIndex].dBufferHead := #TMP_dNextHead;
           #AUX_rgtLastUpdData[#TMP_dIndex] := #INO_tRibbon.rgtGlassData[#TMP_dIndex].rgtBuffer[#TMP_dNextHead];
           #INO_tRibbon.rgtGlassDataUpdate[#TMP_dIndex].xUpdateRequest := FALSE;
       END_IF;

   END_FOR;
END_REGION

REGION Network 6 (SCL): Insert the new glass break or update the last one
   FOR #TMP_dIndex := 0 TO #INO_tRibbon.dActualNumberGlassBreakMachine - 1 DO


       //New position from external device, 
       IF (#INO_tRibbon.rgtGlassBreakUpdate[#TMP_dIndex].xUpdateRequest) THEN

           //Increment the index head
           IF (#INO_tRibbon.rgtGlassBreak[#TMP_dIndex].dBufferHead + 1) >= "DMAXGLASSBREAKSECTORS" THEN
               #TMP_dNextHead := 0;
           ELSE
               #TMP_dNextHead := #INO_tRibbon.rgtGlassBreak[#TMP_dIndex].dBufferHead + 1;
           END_IF;

           //Check if the buffer is full
           IF (#TMP_dNextHead = #INO_tRibbon.rgtGlassBreak[#TMP_dIndex].dBufferTail) AND (#INO_tRibbon.rgtGlassBreak[#TMP_dIndex].dBufferHead <> -1) THEN
               EXIT;
           END_IF; 

           #INO_tRibbon.rgtGlassBreak[#TMP_dIndex].rgtBuffer[#TMP_dNextHead].dEncoderValue_cmm := #INO_tEncoder.dActualEncoderCounter_cmm + #INO_tRibbon.rgtGlassBreak[#TMP_dIndex].dDistSnapRoll_cmm;

           #INO_tRibbon.rgtGlassBreak[#TMP_dIndex].rgtBuffer[#TMP_dNextHead].xGlassBreak := #INO_tRibbon.rgtGlassBreakUpdate[#TMP_dIndex].tData.xGlassBreak;
           #INO_tRibbon.rgtGlassBreak[#TMP_dIndex].rgtBuffer[#TMP_dNextHead].rgxBreakMask := #INO_tRibbon.rgtGlassBreakUpdate[#TMP_dIndex].tData.rgxBreakMask;

           #INO_tRibbon.rgtGlassBreak[#TMP_dIndex].dLastInsertEncCount_cmm := #INO_tRibbon.rgtGlassBreak[#TMP_dIndex].rgtBuffer[#TMP_dNextHead].dEncoderValue_cmm;
           #INO_tRibbon.rgtGlassBreak[#TMP_dIndex].rgtBuffer[#TMP_dNextHead].xUpdateDataBPSA := TRUE;
           #INO_tRibbon.rgtGlassBreak[#TMP_dIndex].rgtBuffer[#TMP_dNextHead].xUpdateDataBPSB := TRUE;
           #INO_tRibbon.rgtGlassBreak[#TMP_dIndex].rgtBuffer[#TMP_dNextHead].xDataPresent := TRUE;

           #INO_tRibbon.rgtGlassBreak[#TMP_dIndex].dBufferHead := #TMP_dNextHead;
           #AUX_rgtLastUpdBreak[#TMP_dIndex] := #INO_tRibbon.rgtGlassBreak[#TMP_dIndex].rgtBuffer[#TMP_dNextHead];
           #INO_tRibbon.rgtGlassBreakUpdate[#TMP_dIndex].xUpdateRequest := FALSE;
       END_IF;

   END_FOR;
END_REGION

REGION Network 7 (SCL): Evaluate glass data request
   FOR #TMP_dIndex := 0 TO "DMAXGLASSDATAREQUEST_IND" DO

       #TMP_dSourceIndex := #INO_tRibbon.rgtGlassDataRequest[#TMP_dIndex].IN_dSourceIndex;

       IF #INO_tRibbon.rgtGlassDataRequest[#TMP_dIndex].IN_xRequestGlassData
           AND NOT #INO_tRibbon.rgtGlassDataRequest[#TMP_dIndex].OUT_xDataReady
           AND #INO_tRibbon.rgtGlassDataRequest[#TMP_dIndex].IN_dSourceIndex < #INO_tRibbon.dActualNumberGlassDataMachine THEN

           //Glass data request, calculate the values. Move data until get less than the distance from user
           #INO_tRibbon.rgtGlassDataRequest[#TMP_dIndex].OUT_dGrossWidth_cmm := #INO_tRibbon.rgtGlassData[#TMP_dSourceIndex].tLastDataBuffer.dGrossWidth_cmm;
           #INO_tRibbon.rgtGlassDataRequest[#TMP_dIndex].OUT_dNetWidth_cmm := #INO_tRibbon.rgtGlassData[#TMP_dSourceIndex].tLastDataBuffer.dNetWidth_cmm;
           #INO_tRibbon.rgtGlassDataRequest[#TMP_dIndex].OUT_dGrossWander_cmm := #INO_tRibbon.rgtGlassData[#TMP_dSourceIndex].tLastDataBuffer.dGrossWander_cmm;
           #INO_tRibbon.rgtGlassDataRequest[#TMP_dIndex].OUT_dNetWander_cmm := #INO_tRibbon.rgtGlassData[#TMP_dSourceIndex].tLastDataBuffer.dNetWander_cmm;

           #TMP_dNextTail := #INO_tRibbon.rgtGlassData[#TMP_dSourceIndex].dBufferTail;

           WHILE (#TMP_dNextTail <> #INO_tRibbon.rgtGlassData[#TMP_dSourceIndex].dBufferHead)
               AND (#INO_tRibbon.rgtGlassData[#TMP_dSourceIndex].dBufferHead <> -1) DO

